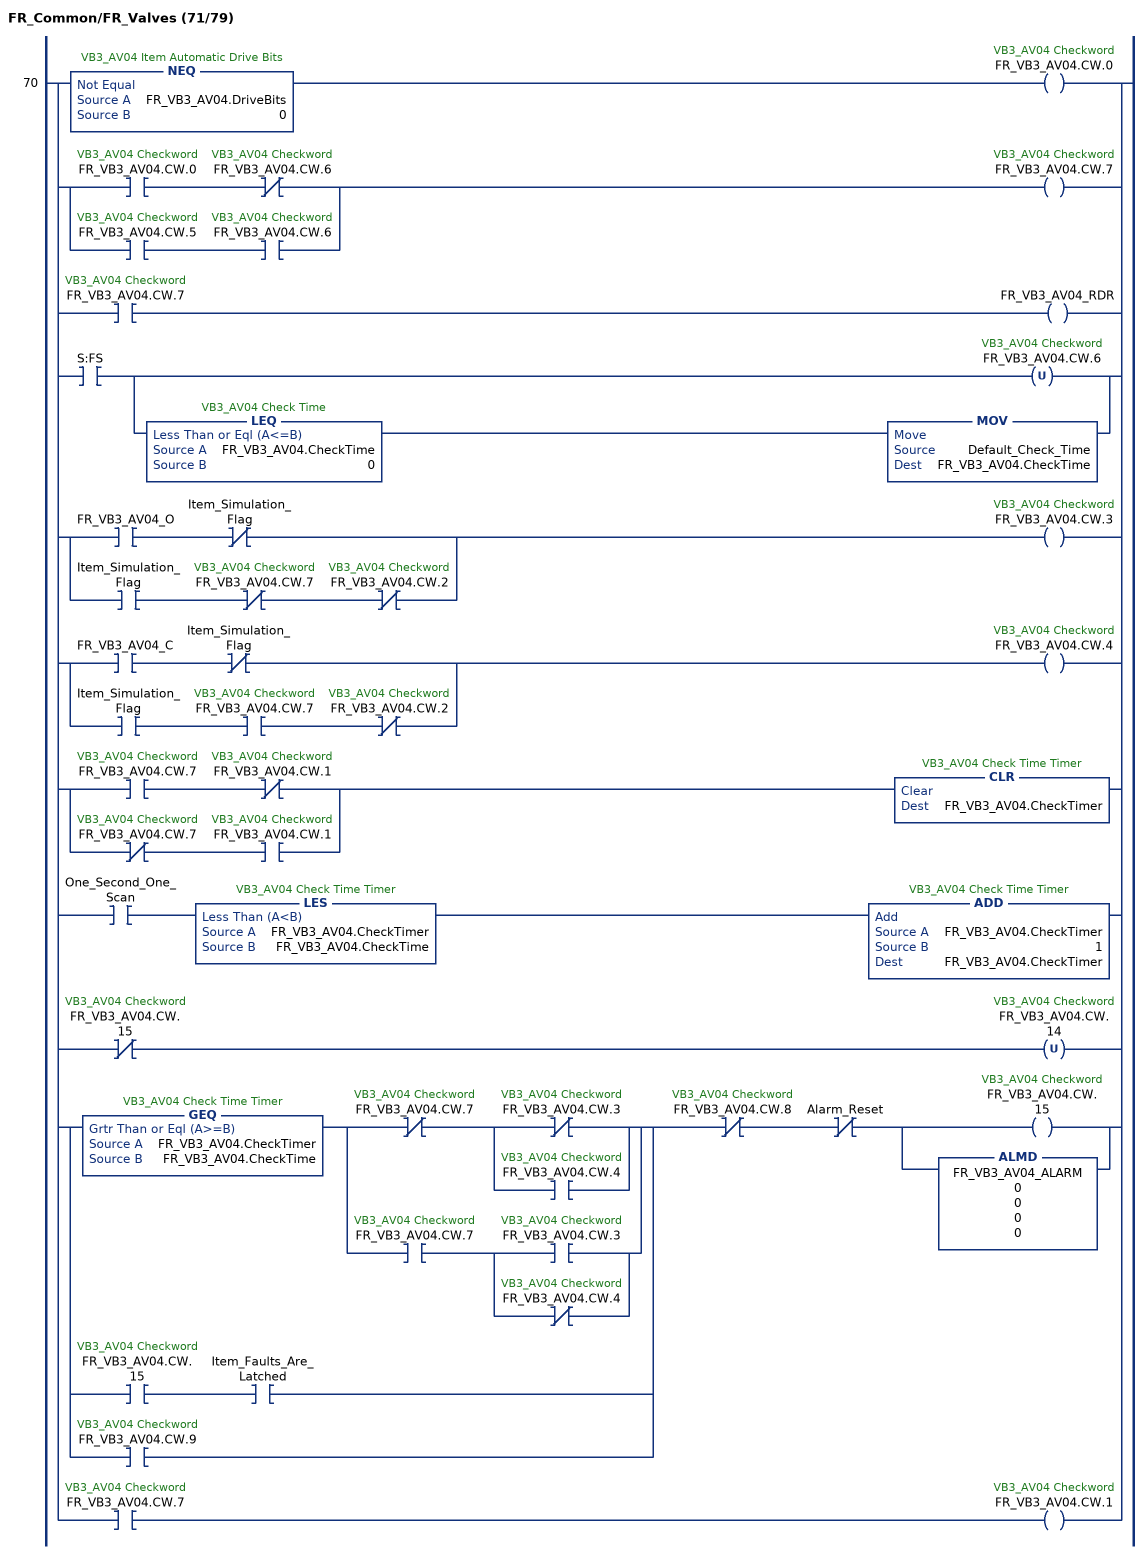
   70: [NEQ(FR_VB3_AV04.DriveBits,0) OTE(FR_VB3_AV04.CW.0) ,[XIC(FR_VB3_AV04.CW.0) XIO(FR_VB3_AV04.CW.6) ,XIC(FR_VB3_AV04.CW.5) XIC(FR_VB3_AV04.CW.6) ] OTE(FR_VB3_AV04.CW.7) ,XIC(FR_VB3_AV04.CW.7) OTE(FR_VB3_AV04_RDR) ,XIC(S:FS) [OTU(FR_VB3_AV04.CW.6) ,LEQ(FR_VB3_AV04.CheckTime,0) MOV(Default_Check_Time,FR_VB3_AV04.CheckTime) ] ,[[XIC(FR_VB3_AV04_O) XIO(Item_Simulation_Flag) ,XIC(Item_Simulation_Flag) XIO(FR_VB3_AV04.CW.7) XIO(FR_VB3_AV04.CW.2) ] OTE(FR_VB3_AV04.CW.3) ,[XIC(FR_VB3_AV04_C) XIO(Item_Simulation_Flag) ,XIC(Item_Simulation_Flag) XIC(FR_VB3_AV04.CW.7) XIO(FR_VB3_AV04.CW.2) ] OTE(FR_VB3_AV04.CW.4) ] ,[XIC(FR_VB3_AV04.CW.7) XIO(FR_VB3_AV04.CW.1) ,XIO(FR_VB3_AV04.CW.7) XIC(FR_VB3_AV04.CW.1) ] CLR(FR_VB3_AV04.CheckTimer) ,XIC(One_Second_One_Scan) LES(FR_VB3_AV04.CheckTimer,FR_VB3_AV04.CheckTime) ADD(FR_VB3_AV04.CheckTimer,1,FR_VB3_AV04.CheckTimer) ,XIO(FR_VB3_AV04.CW.15) OTU(FR_VB3_AV04.CW.14) ,[GEQ(FR_VB3_AV04.CheckTimer,FR_VB3_AV04.CheckTime) [XIO(FR_VB3_AV04.CW.7) [XIO(FR_VB3_AV04.CW.3) ,XIC(FR_VB3_AV04.CW.4) ] ,XIC(FR_VB3_AV04.CW.7) [XIC(FR_VB3_AV04.CW.3) ,XIO(FR_VB3_AV04.CW.4) ] ] ,XIC(FR_VB3_AV04.CW.15) XIC(Item_Faults_Are_Latched) ,XIC(FR_VB3_AV04.CW.9) ] XIO(FR_VB3_AV04.CW.8) XIO(Alarm_Reset) [OTE(FR_VB3_AV04.CW.15) ,ALMD(FR_VB3_AV04_ALARM,0,0,0,0) ] ,XIC(FR_VB3_AV04.CW.7) OTE(FR_VB3_AV04.CW.1) ];
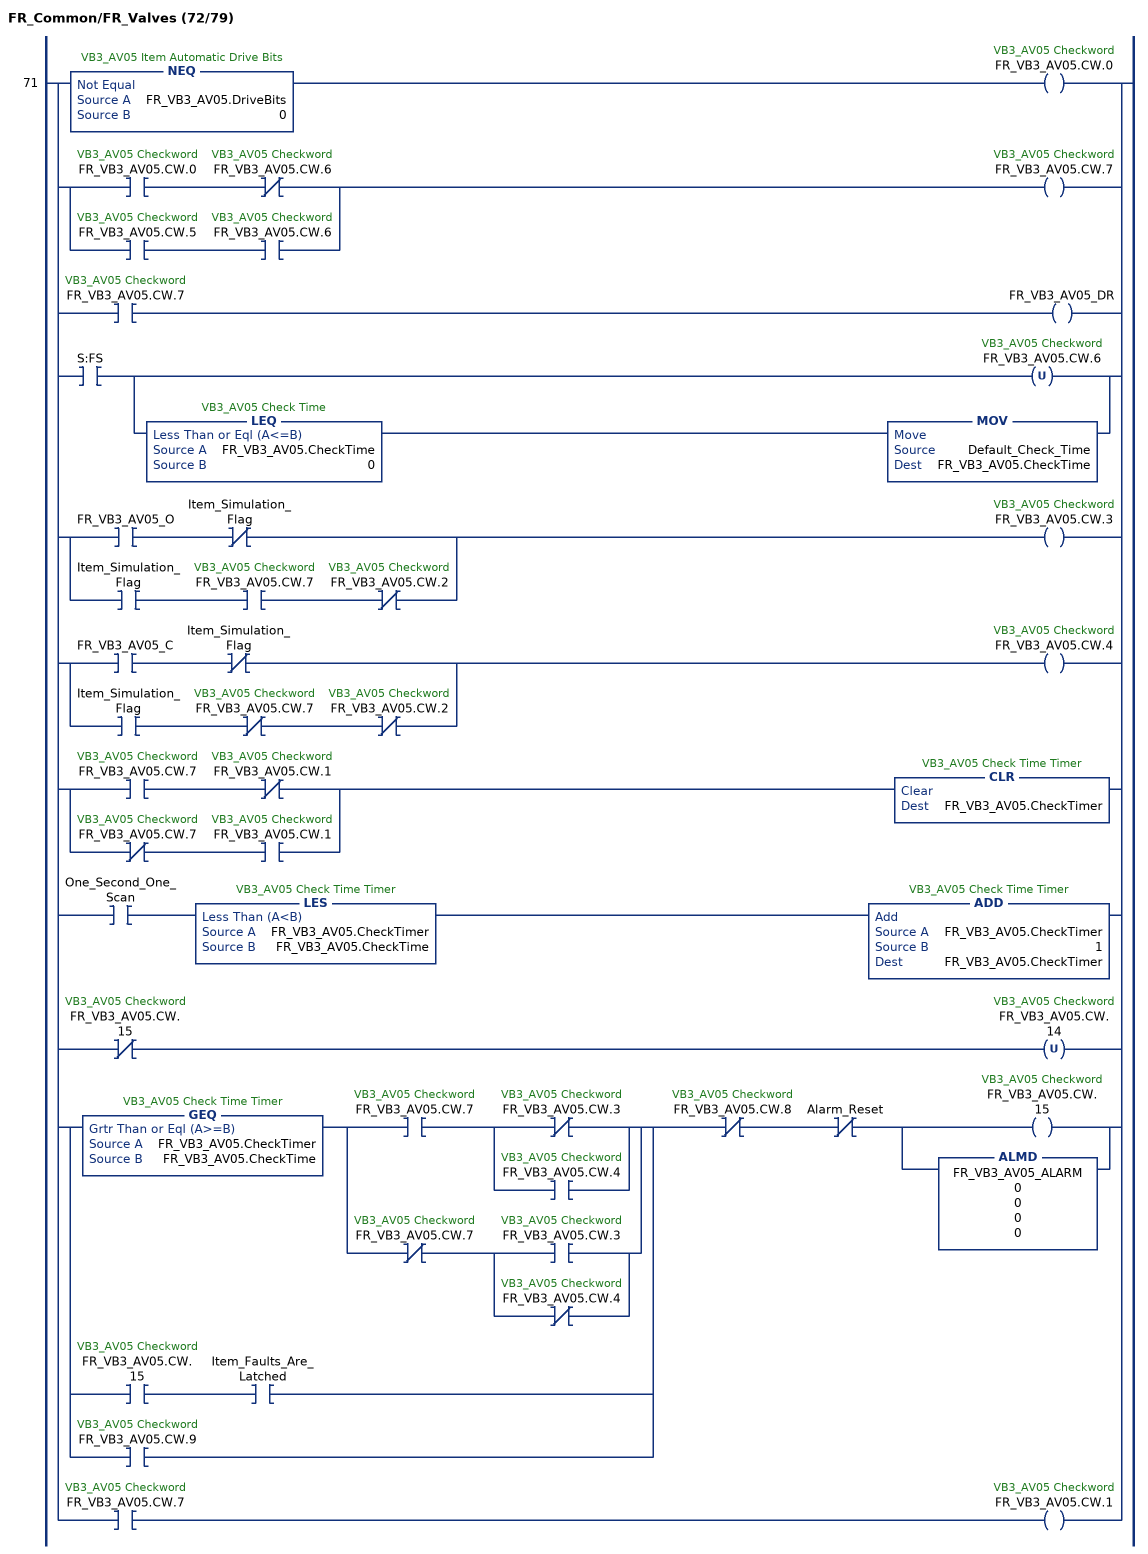
   71: [NEQ(FR_VB3_AV05.DriveBits,0) OTE(FR_VB3_AV05.CW.0) ,[XIC(FR_VB3_AV05.CW.0) XIO(FR_VB3_AV05.CW.6) ,XIC(FR_VB3_AV05.CW.5) XIC(FR_VB3_AV05.CW.6) ] OTE(FR_VB3_AV05.CW.7) ,XIC(FR_VB3_AV05.CW.7) OTE(FR_VB3_AV05_DR) ,XIC(S:FS) [OTU(FR_VB3_AV05.CW.6) ,LEQ(FR_VB3_AV05.CheckTime,0) MOV(Default_Check_Time,FR_VB3_AV05.CheckTime) ] ,[[XIC(FR_VB3_AV05_O) XIO(Item_Simulation_Flag) ,XIC(Item_Simulation_Flag) XIC(FR_VB3_AV05.CW.7) XIO(FR_VB3_AV05.CW.2) ] OTE(FR_VB3_AV05.CW.3) ,[XIC(FR_VB3_AV05_C) XIO(Item_Simulation_Flag) ,XIC(Item_Simulation_Flag) XIO(FR_VB3_AV05.CW.7) XIO(FR_VB3_AV05.CW.2) ] OTE(FR_VB3_AV05.CW.4) ] ,[XIC(FR_VB3_AV05.CW.7) XIO(FR_VB3_AV05.CW.1) ,XIO(FR_VB3_AV05.CW.7) XIC(FR_VB3_AV05.CW.1) ] CLR(FR_VB3_AV05.CheckTimer) ,XIC(One_Second_One_Scan) LES(FR_VB3_AV05.CheckTimer,FR_VB3_AV05.CheckTime) ADD(FR_VB3_AV05.CheckTimer,1,FR_VB3_AV05.CheckTimer) ,XIO(FR_VB3_AV05.CW.15) OTU(FR_VB3_AV05.CW.14) ,[GEQ(FR_VB3_AV05.CheckTimer,FR_VB3_AV05.CheckTime) [XIC(FR_VB3_AV05.CW.7) [XIO(FR_VB3_AV05.CW.3) ,XIC(FR_VB3_AV05.CW.4) ] ,XIO(FR_VB3_AV05.CW.7) [XIC(FR_VB3_AV05.CW.3) ,XIO(FR_VB3_AV05.CW.4) ] ] ,XIC(FR_VB3_AV05.CW.15) XIC(Item_Faults_Are_Latched) ,XIC(FR_VB3_AV05.CW.9) ] XIO(FR_VB3_AV05.CW.8) XIO(Alarm_Reset) [OTE(FR_VB3_AV05.CW.15) ,ALMD(FR_VB3_AV05_ALARM,0,0,0,0) ] ,XIC(FR_VB3_AV05.CW.7) OTE(FR_VB3_AV05.CW.1) ];
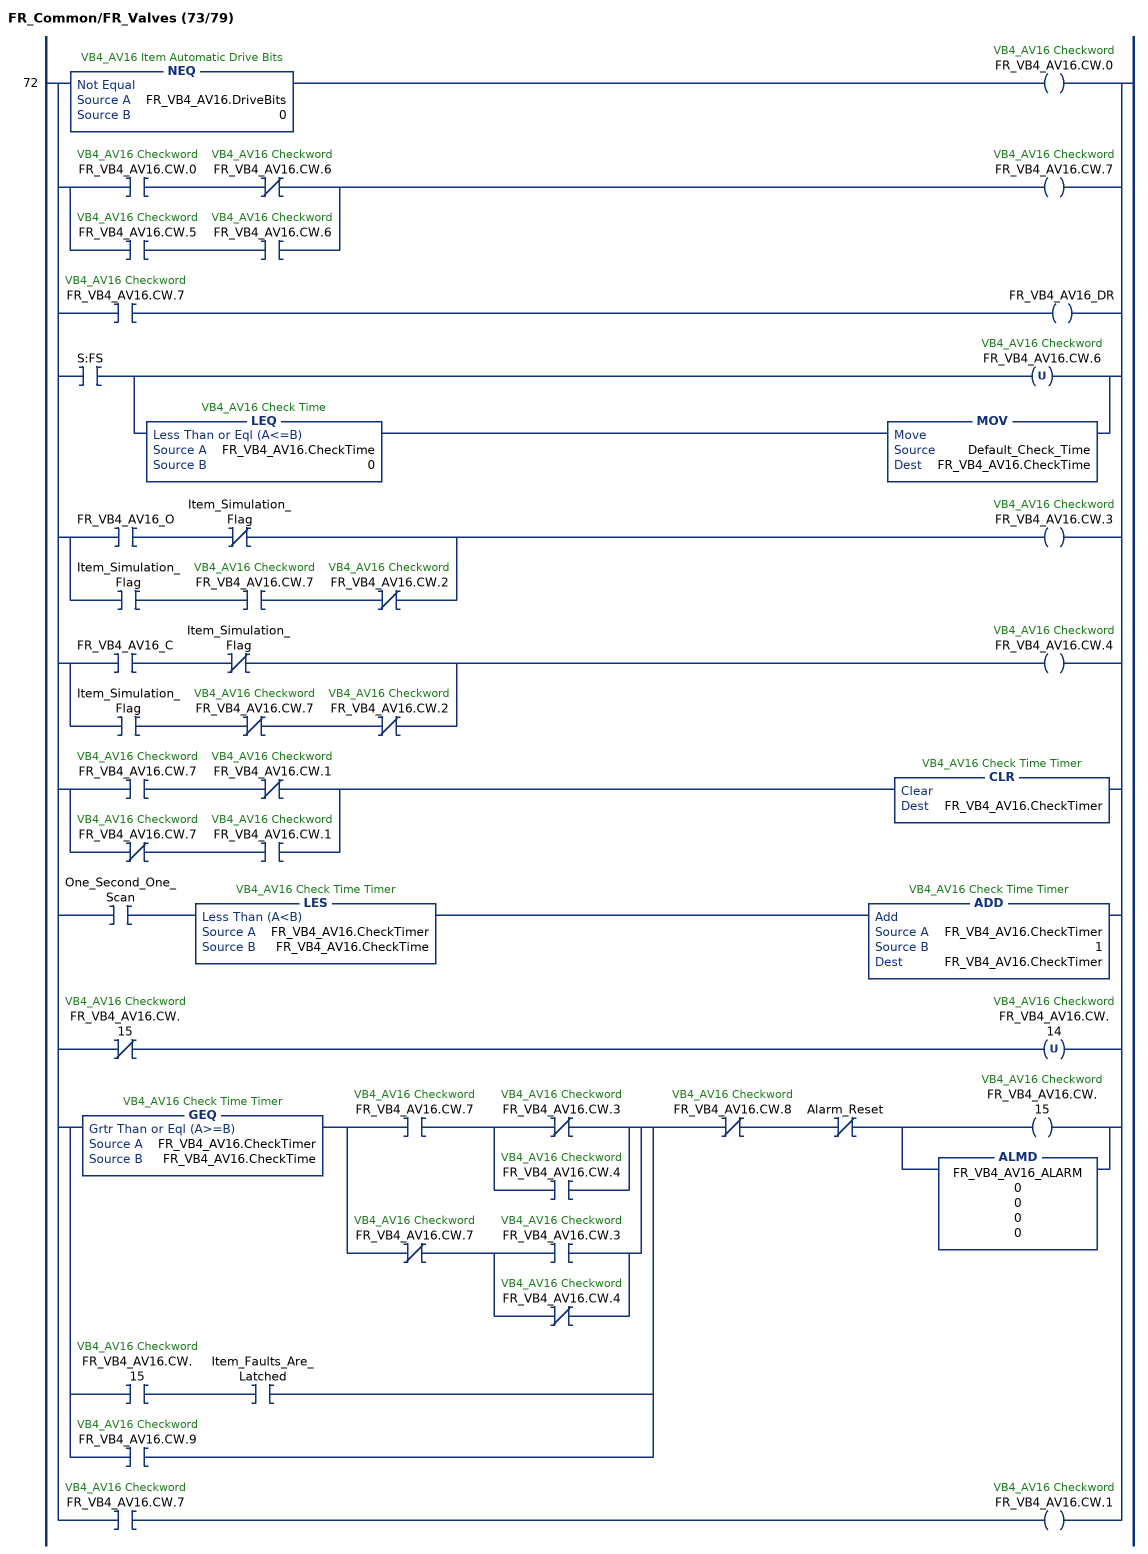
   72: [NEQ(FR_VB4_AV16.DriveBits,0) OTE(FR_VB4_AV16.CW.0) ,[XIC(FR_VB4_AV16.CW.0) XIO(FR_VB4_AV16.CW.6) ,XIC(FR_VB4_AV16.CW.5) XIC(FR_VB4_AV16.CW.6) ] OTE(FR_VB4_AV16.CW.7) ,XIC(FR_VB4_AV16.CW.7) OTE(FR_VB4_AV16_DR) ,XIC(S:FS) [OTU(FR_VB4_AV16.CW.6) ,LEQ(FR_VB4_AV16.CheckTime,0) MOV(Default_Check_Time,FR_VB4_AV16.CheckTime) ] ,[[XIC(FR_VB4_AV16_O) XIO(Item_Simulation_Flag) ,XIC(Item_Simulation_Flag) XIC(FR_VB4_AV16.CW.7) XIO(FR_VB4_AV16.CW.2) ] OTE(FR_VB4_AV16.CW.3) ,[XIC(FR_VB4_AV16_C) XIO(Item_Simulation_Flag) ,XIC(Item_Simulation_Flag) XIO(FR_VB4_AV16.CW.7) XIO(FR_VB4_AV16.CW.2) ] OTE(FR_VB4_AV16.CW.4) ] ,[XIC(FR_VB4_AV16.CW.7) XIO(FR_VB4_AV16.CW.1) ,XIO(FR_VB4_AV16.CW.7) XIC(FR_VB4_AV16.CW.1) ] CLR(FR_VB4_AV16.CheckTimer) ,XIC(One_Second_One_Scan) LES(FR_VB4_AV16.CheckTimer,FR_VB4_AV16.CheckTime) ADD(FR_VB4_AV16.CheckTimer,1,FR_VB4_AV16.CheckTimer) ,XIO(FR_VB4_AV16.CW.15) OTU(FR_VB4_AV16.CW.14) ,[GEQ(FR_VB4_AV16.CheckTimer,FR_VB4_AV16.CheckTime) [XIC(FR_VB4_AV16.CW.7) [XIO(FR_VB4_AV16.CW.3) ,XIC(FR_VB4_AV16.CW.4) ] ,XIO(FR_VB4_AV16.CW.7) [XIC(FR_VB4_AV16.CW.3) ,XIO(FR_VB4_AV16.CW.4) ] ] ,XIC(FR_VB4_AV16.CW.15) XIC(Item_Faults_Are_Latched) ,XIC(FR_VB4_AV16.CW.9) ] XIO(FR_VB4_AV16.CW.8) XIO(Alarm_Reset) [OTE(FR_VB4_AV16.CW.15) ,ALMD(FR_VB4_AV16_ALARM,0,0,0,0) ] ,XIC(FR_VB4_AV16.CW.7) OTE(FR_VB4_AV16.CW.1) ];
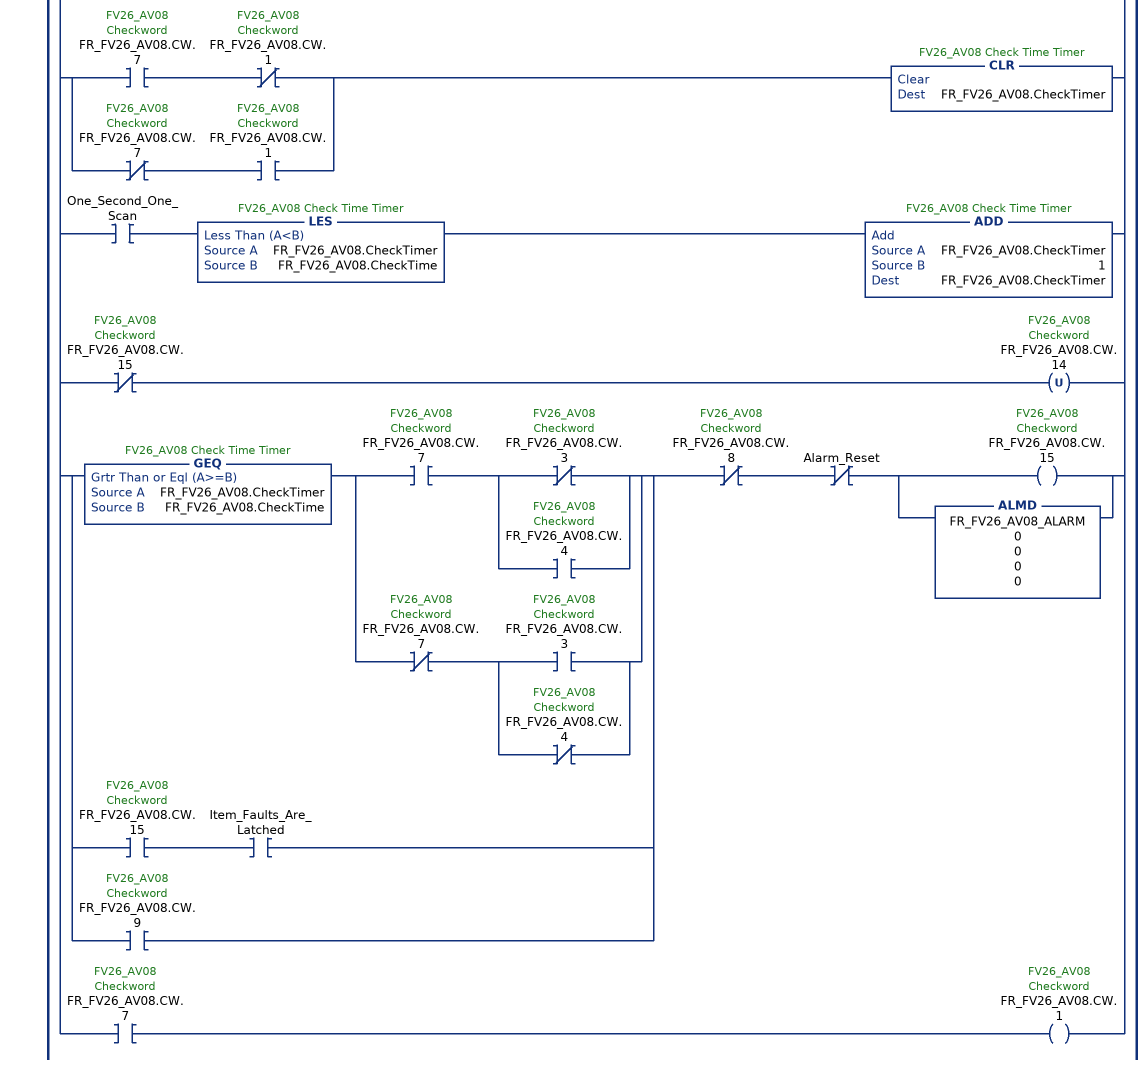
   73: [NEQ(FR_FV26_AV08.DriveBits,0) OTE(FR_FV26_AV08.CW.0) ,[XIC(FR_FV26_AV08.CW.0) XIO(FR_FV26_AV08.CW.6) ,XIC(FR_FV26_AV08.CW.5) XIC(FR_FV26_AV08.CW.6) ] OTE(FR_FV26_AV08.CW.7) ,XIC(FR_FV26_AV08.CW.7) OTE(FR_FV26_AV08_DR) ,XIC(S:FS) [OTU(FR_FV26_AV08.CW.6) ,LEQ(FR_FV26_AV08.CheckTime,0) MOV(Default_Check_Time,FR_FV26_AV08.CheckTime) ] ,[[XIC(FR_FV26_AV08_O) XIO(Item_Simulation_Flag) ,XIC(Item_Simulation_Flag) XIC(FR_FV26_AV08.CW.7) XIO(FR_FV26_AV08.CW.2) ] OTE(FR_FV26_AV08.CW.3) ,[XIC(FR_FV26_AV08_C) XIO(Item_Simulation_Flag) ,XIC(Item_Simulation_Flag) XIO(FR_FV26_AV08.CW.7) XIO(FR_FV26_AV08.CW.2) ] OTE(FR_FV26_AV08.CW.4) ] ,[XIC(FR_FV26_AV08.CW.7) XIO(FR_FV26_AV08.CW.1) ,XIO(FR_FV26_AV08.CW.7) XIC(FR_FV26_AV08.CW.1) ] CLR(FR_FV26_AV08.CheckTimer) ,XIC(One_Second_One_Scan) LES(FR_FV26_AV08.CheckTimer,FR_FV26_AV08.CheckTime) ADD(FR_FV26_AV08.CheckTimer,1,FR_FV26_AV08.CheckTimer) ,XIO(FR_FV26_AV08.CW.15) OTU(FR_FV26_AV08.CW.14) ,[GEQ(FR_FV26_AV08.CheckTimer,FR_FV26_AV08.CheckTime) [XIC(FR_FV26_AV08.CW.7) [XIO(FR_FV26_AV08.CW.3) ,XIC(FR_FV26_AV08.CW.4) ] ,XIO(FR_FV26_AV08.CW.7) [XIC(FR_FV26_AV08.CW.3) ,XIO(FR_FV26_AV08.CW.4) ] ] ,XIC(FR_FV26_AV08.CW.15) XIC(Item_Faults_Are_Latched) ,XIC(FR_FV26_AV08.CW.9) ] XIO(FR_FV26_AV08.CW.8) XIO(Alarm_Reset) [OTE(FR_FV26_AV08.CW.15) ,ALMD(FR_FV26_AV08_ALARM,0,0,0,0) ] ,XIC(FR_FV26_AV08.CW.7) OTE(FR_FV26_AV08.CW.1) ];
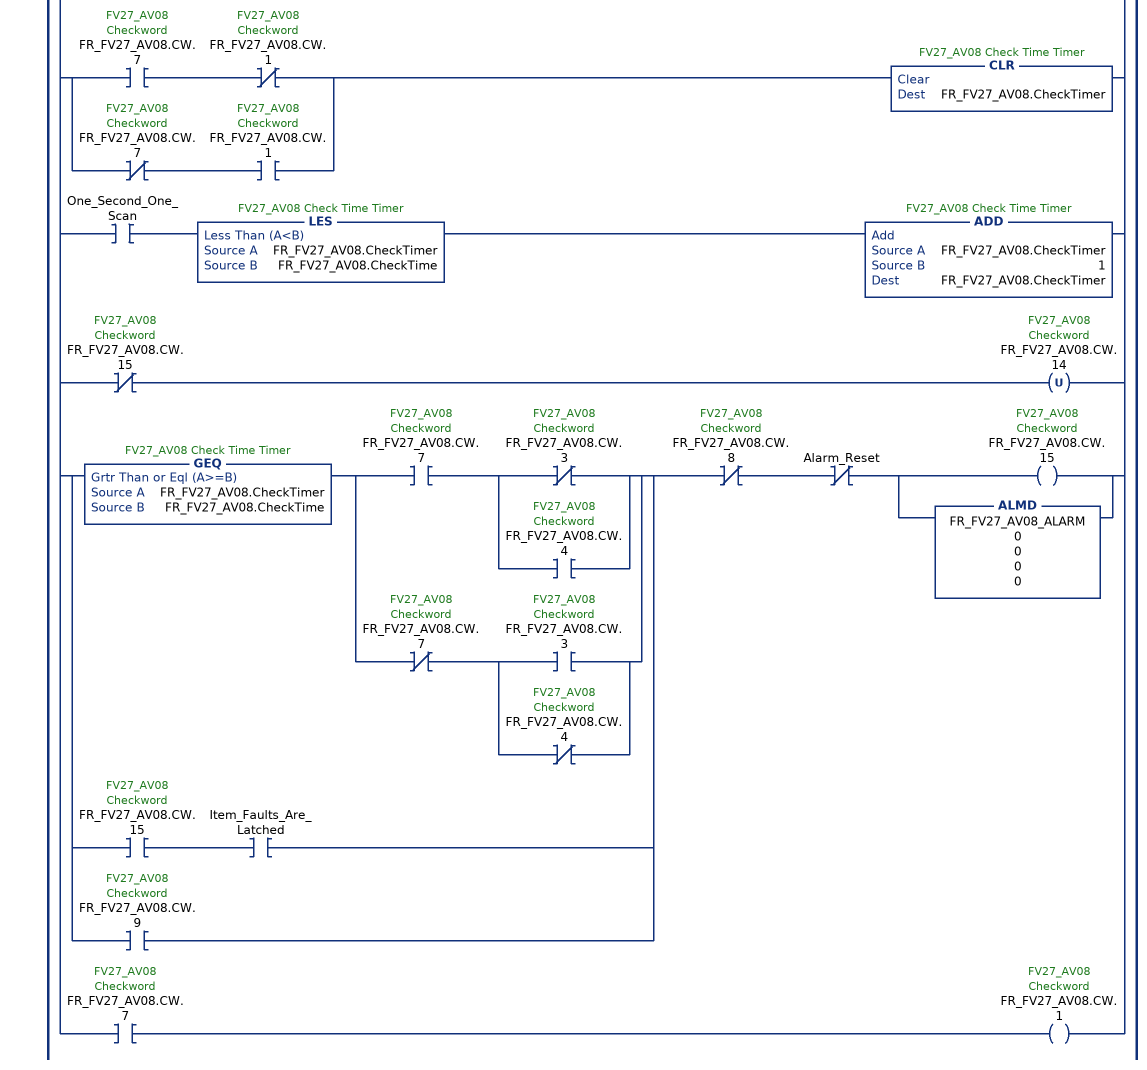
   74: [NEQ(FR_FV27_AV08.DriveBits,0) OTE(FR_FV27_AV08.CW.0) ,[XIC(FR_FV27_AV08.CW.0) XIO(FR_FV27_AV08.CW.6) ,XIC(FR_FV27_AV08.CW.5) XIC(FR_FV27_AV08.CW.6) ] OTE(FR_FV27_AV08.CW.7) ,XIC(FR_FV27_AV08.CW.7) OTE(FR_FV27_AV08_DR) ,XIC(S:FS) [OTU(FR_FV27_AV08.CW.6) ,LEQ(FR_FV27_AV08.CheckTime,0) MOV(Default_Check_Time,FR_FV27_AV08.CheckTime) ] ,[[XIC(FR_FV27_AV08_O) XIO(Item_Simulation_Flag) ,XIC(Item_Simulation_Flag) XIC(FR_FV27_AV08.CW.7) XIO(FR_FV27_AV08.CW.2) ] OTE(FR_FV27_AV08.CW.3) ,[XIC(FR_FV27_AV08_C) XIO(Item_Simulation_Flag) ,XIC(Item_Simulation_Flag) XIO(FR_FV27_AV08.CW.7) XIO(FR_FV27_AV08.CW.2) ] OTE(FR_FV27_AV08.CW.4) ] ,[XIC(FR_FV27_AV08.CW.7) XIO(FR_FV27_AV08.CW.1) ,XIO(FR_FV27_AV08.CW.7) XIC(FR_FV27_AV08.CW.1) ] CLR(FR_FV27_AV08.CheckTimer) ,XIC(One_Second_One_Scan) LES(FR_FV27_AV08.CheckTimer,FR_FV27_AV08.CheckTime) ADD(FR_FV27_AV08.CheckTimer,1,FR_FV27_AV08.CheckTimer) ,XIO(FR_FV27_AV08.CW.15) OTU(FR_FV27_AV08.CW.14) ,[GEQ(FR_FV27_AV08.CheckTimer,FR_FV27_AV08.CheckTime) [XIC(FR_FV27_AV08.CW.7) [XIO(FR_FV27_AV08.CW.3) ,XIC(FR_FV27_AV08.CW.4) ] ,XIO(FR_FV27_AV08.CW.7) [XIC(FR_FV27_AV08.CW.3) ,XIO(FR_FV27_AV08.CW.4) ] ] ,XIC(FR_FV27_AV08.CW.15) XIC(Item_Faults_Are_Latched) ,XIC(FR_FV27_AV08.CW.9) ] XIO(FR_FV27_AV08.CW.8) XIO(Alarm_Reset) [OTE(FR_FV27_AV08.CW.15) ,ALMD(FR_FV27_AV08_ALARM,0,0,0,0) ] ,XIC(FR_FV27_AV08.CW.7) OTE(FR_FV27_AV08.CW.1) ];
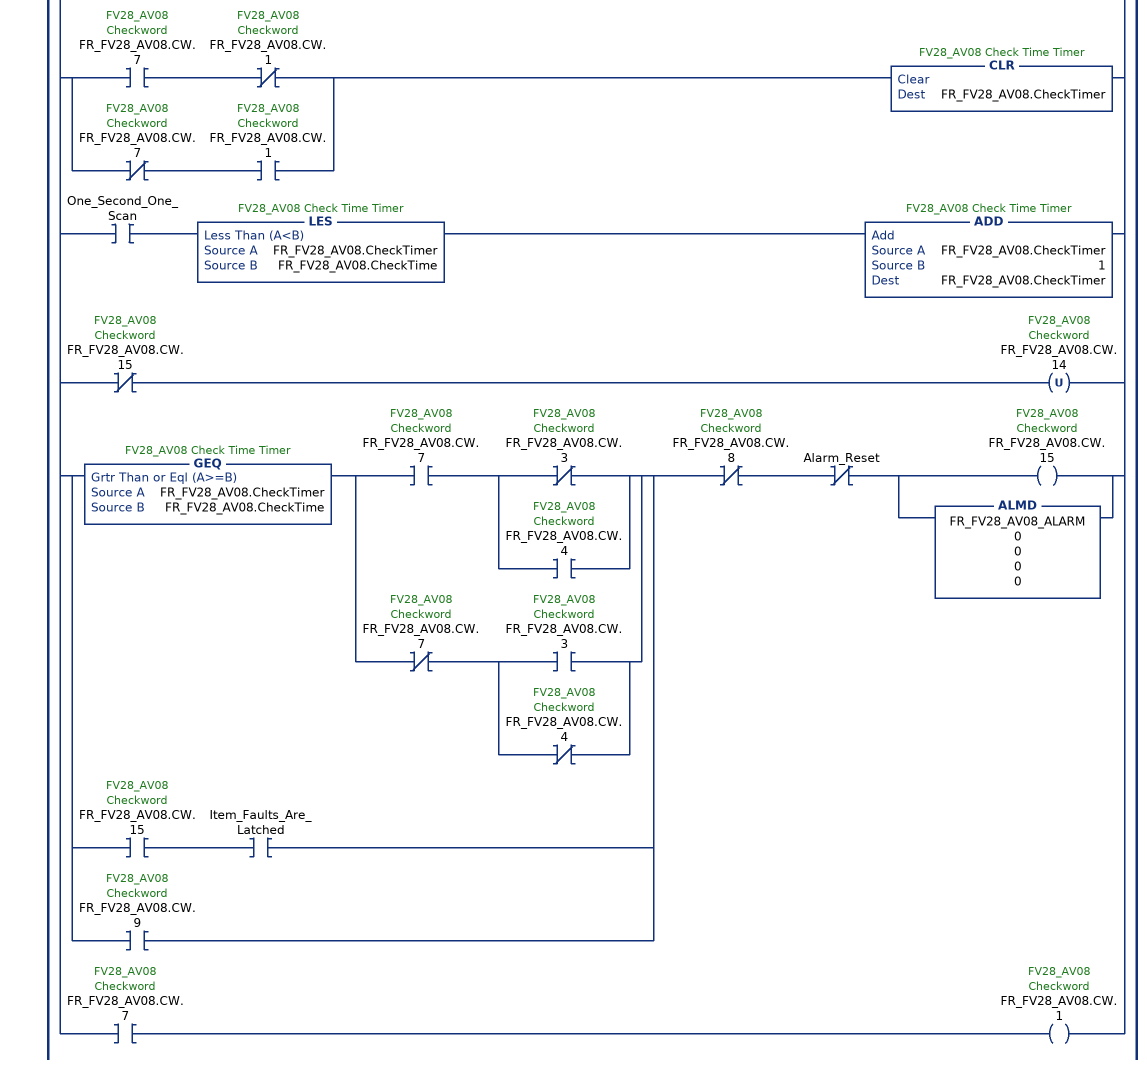
   75: [NEQ(FR_FV28_AV08.DriveBits,0) OTE(FR_FV28_AV08.CW.0) ,[XIC(FR_FV28_AV08.CW.0) XIO(FR_FV28_AV08.CW.6) ,XIC(FR_FV28_AV08.CW.5) XIC(FR_FV28_AV08.CW.6) ] OTE(FR_FV28_AV08.CW.7) ,XIC(FR_FV28_AV08.CW.7) OTE(FR_FV28_AV08_DR) ,XIC(S:FS) [OTU(FR_FV28_AV08.CW.6) ,LEQ(FR_FV28_AV08.CheckTime,0) MOV(Default_Check_Time,FR_FV28_AV08.CheckTime) ] ,[[XIC(FR_FV28_AV08_O) XIO(Item_Simulation_Flag) ,XIC(Item_Simulation_Flag) XIC(FR_FV28_AV08.CW.7) XIO(FR_FV28_AV08.CW.2) ] OTE(FR_FV28_AV08.CW.3) ,[XIC(FR_FV28_AV08_C) XIO(Item_Simulation_Flag) ,XIC(Item_Simulation_Flag) XIO(FR_FV28_AV08.CW.7) XIO(FR_FV28_AV08.CW.2) ] OTE(FR_FV28_AV08.CW.4) ] ,[XIC(FR_FV28_AV08.CW.7) XIO(FR_FV28_AV08.CW.1) ,XIO(FR_FV28_AV08.CW.7) XIC(FR_FV28_AV08.CW.1) ] CLR(FR_FV28_AV08.CheckTimer) ,XIC(One_Second_One_Scan) LES(FR_FV28_AV08.CheckTimer,FR_FV28_AV08.CheckTime) ADD(FR_FV28_AV08.CheckTimer,1,FR_FV28_AV08.CheckTimer) ,XIO(FR_FV28_AV08.CW.15) OTU(FR_FV28_AV08.CW.14) ,[GEQ(FR_FV28_AV08.CheckTimer,FR_FV28_AV08.CheckTime) [XIC(FR_FV28_AV08.CW.7) [XIO(FR_FV28_AV08.CW.3) ,XIC(FR_FV28_AV08.CW.4) ] ,XIO(FR_FV28_AV08.CW.7) [XIC(FR_FV28_AV08.CW.3) ,XIO(FR_FV28_AV08.CW.4) ] ] ,XIC(FR_FV28_AV08.CW.15) XIC(Item_Faults_Are_Latched) ,XIC(FR_FV28_AV08.CW.9) ] XIO(FR_FV28_AV08.CW.8) XIO(Alarm_Reset) [OTE(FR_FV28_AV08.CW.15) ,ALMD(FR_FV28_AV08_ALARM,0,0,0,0) ] ,XIC(FR_FV28_AV08.CW.7) OTE(FR_FV28_AV08.CW.1) ];
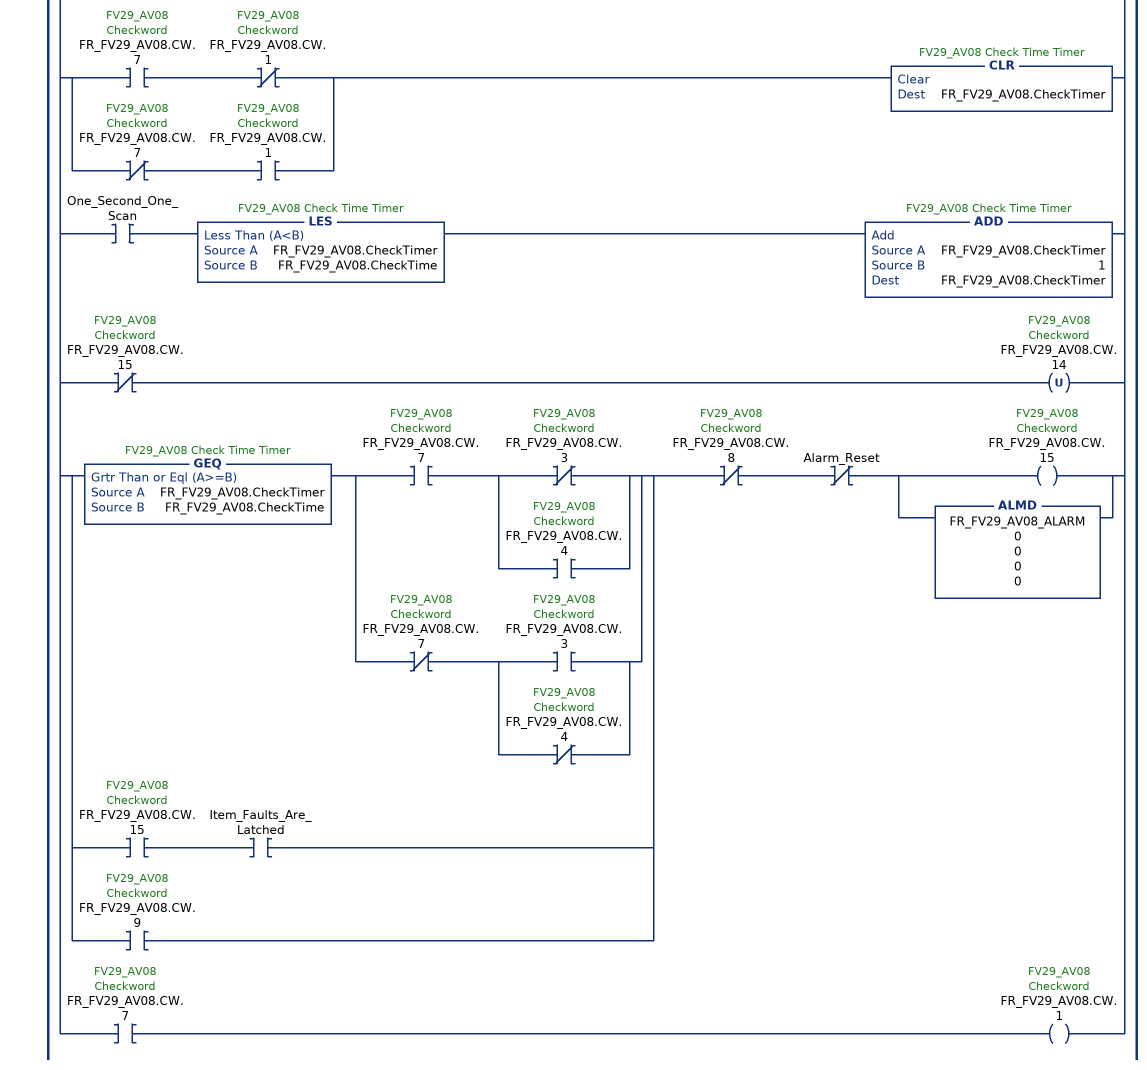
   76: [NEQ(FR_FV29_AV08.DriveBits,0) OTE(FR_FV29_AV08.CW.0) ,[XIC(FR_FV29_AV08.CW.0) XIO(FR_FV29_AV08.CW.6) ,XIC(FR_FV29_AV08.CW.5) XIC(FR_FV29_AV08.CW.6) ] OTE(FR_FV29_AV08.CW.7) ,XIC(FR_FV29_AV08.CW.7) OTE(FR_FV29_AV08_DR) ,XIC(S:FS) [OTU(FR_FV29_AV08.CW.6) ,LEQ(FR_FV29_AV08.CheckTime,0) MOV(Default_Check_Time,FR_FV29_AV08.CheckTime) ] ,[[XIC(FR_FV29_AV08_O) XIO(Item_Simulation_Flag) ,XIC(Item_Simulation_Flag) XIC(FR_FV29_AV08.CW.7) XIO(FR_FV29_AV08.CW.2) ] OTE(FR_FV29_AV08.CW.3) ,[XIC(FR_FV29_AV08_C) XIO(Item_Simulation_Flag) ,XIC(Item_Simulation_Flag) XIO(FR_FV29_AV08.CW.7) XIO(FR_FV29_AV08.CW.2) ] OTE(FR_FV29_AV08.CW.4) ] ,[XIC(FR_FV29_AV08.CW.7) XIO(FR_FV29_AV08.CW.1) ,XIO(FR_FV29_AV08.CW.7) XIC(FR_FV29_AV08.CW.1) ] CLR(FR_FV29_AV08.CheckTimer) ,XIC(One_Second_One_Scan) LES(FR_FV29_AV08.CheckTimer,FR_FV29_AV08.CheckTime) ADD(FR_FV29_AV08.CheckTimer,1,FR_FV29_AV08.CheckTimer) ,XIO(FR_FV29_AV08.CW.15) OTU(FR_FV29_AV08.CW.14) ,[GEQ(FR_FV29_AV08.CheckTimer,FR_FV29_AV08.CheckTime) [XIC(FR_FV29_AV08.CW.7) [XIO(FR_FV29_AV08.CW.3) ,XIC(FR_FV29_AV08.CW.4) ] ,XIO(FR_FV29_AV08.CW.7) [XIC(FR_FV29_AV08.CW.3) ,XIO(FR_FV29_AV08.CW.4) ] ] ,XIC(FR_FV29_AV08.CW.15) XIC(Item_Faults_Are_Latched) ,XIC(FR_FV29_AV08.CW.9) ] XIO(FR_FV29_AV08.CW.8) XIO(Alarm_Reset) [OTE(FR_FV29_AV08.CW.15) ,ALMD(FR_FV29_AV08_ALARM,0,0,0,0) ] ,XIC(FR_FV29_AV08.CW.7) OTE(FR_FV29_AV08.CW.1) ];
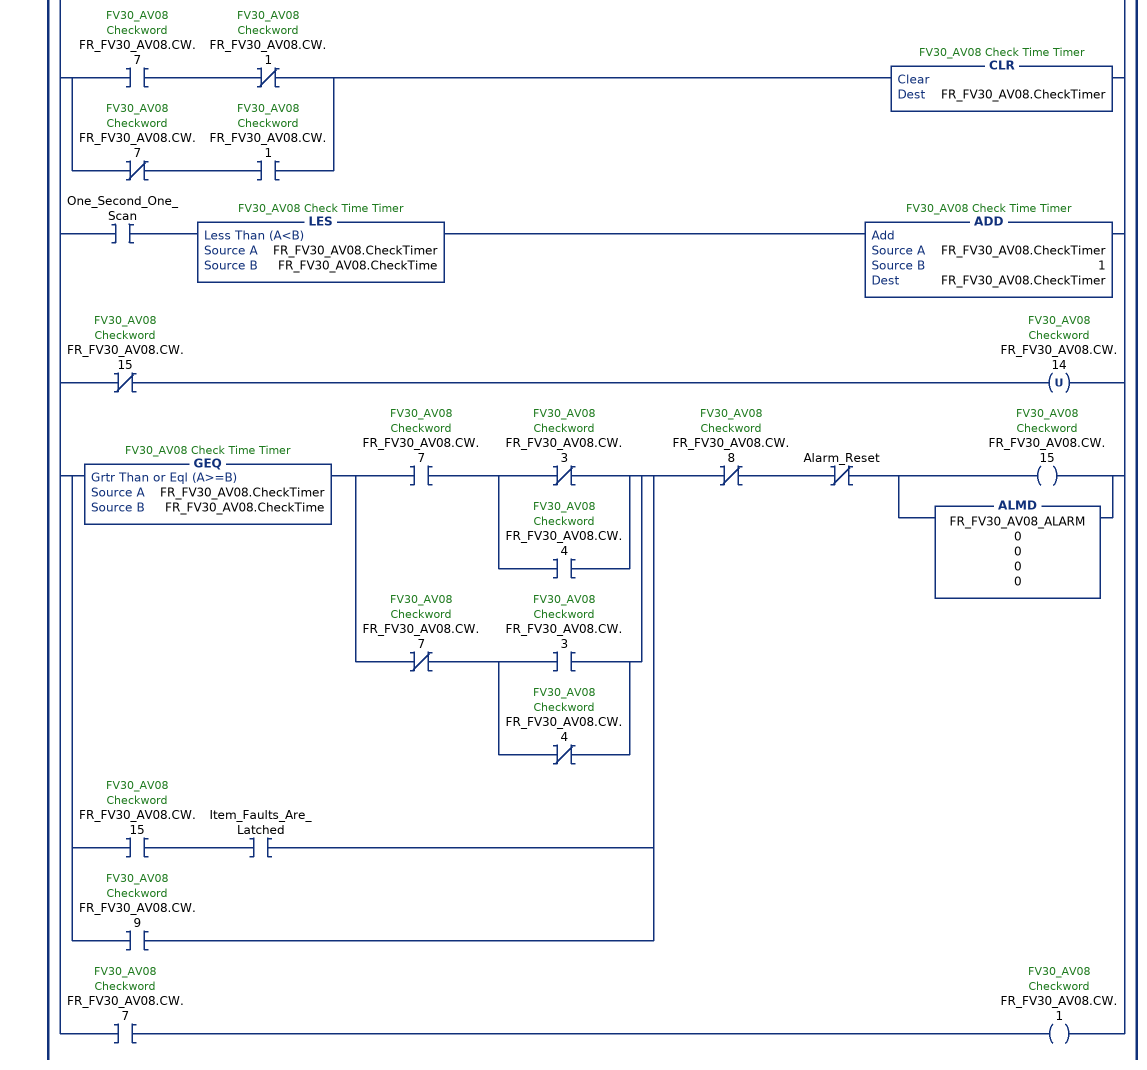
   77: [NEQ(FR_FV30_AV08.DriveBits,0) OTE(FR_FV30_AV08.CW.0) ,[XIC(FR_FV30_AV08.CW.0) XIO(FR_FV30_AV08.CW.6) ,XIC(FR_FV30_AV08.CW.5) XIC(FR_FV30_AV08.CW.6) ] OTE(FR_FV30_AV08.CW.7) ,XIC(FR_FV30_AV08.CW.7) OTE(FR_FV30_AV08_DR) ,XIC(S:FS) [OTU(FR_FV30_AV08.CW.6) ,LEQ(FR_FV30_AV08.CheckTime,0) MOV(Default_Check_Time,FR_FV30_AV08.CheckTime) ] ,[[XIC(FR_FV30_AV08_O) XIO(Item_Simulation_Flag) ,XIC(Item_Simulation_Flag) XIC(FR_FV30_AV08.CW.7) XIO(FR_FV30_AV08.CW.2) ] OTE(FR_FV30_AV08.CW.3) ,[XIC(FR_FV30_AV08_C) XIO(Item_Simulation_Flag) ,XIC(Item_Simulation_Flag) XIO(FR_FV30_AV08.CW.7) XIO(FR_FV30_AV08.CW.2) ] OTE(FR_FV30_AV08.CW.4) ] ,[XIC(FR_FV30_AV08.CW.7) XIO(FR_FV30_AV08.CW.1) ,XIO(FR_FV30_AV08.CW.7) XIC(FR_FV30_AV08.CW.1) ] CLR(FR_FV30_AV08.CheckTimer) ,XIC(One_Second_One_Scan) LES(FR_FV30_AV08.CheckTimer,FR_FV30_AV08.CheckTime) ADD(FR_FV30_AV08.CheckTimer,1,FR_FV30_AV08.CheckTimer) ,XIO(FR_FV30_AV08.CW.15) OTU(FR_FV30_AV08.CW.14) ,[GEQ(FR_FV30_AV08.CheckTimer,FR_FV30_AV08.CheckTime) [XIC(FR_FV30_AV08.CW.7) [XIO(FR_FV30_AV08.CW.3) ,XIC(FR_FV30_AV08.CW.4) ] ,XIO(FR_FV30_AV08.CW.7) [XIC(FR_FV30_AV08.CW.3) ,XIO(FR_FV30_AV08.CW.4) ] ] ,XIC(FR_FV30_AV08.CW.15) XIC(Item_Faults_Are_Latched) ,XIC(FR_FV30_AV08.CW.9) ] XIO(FR_FV30_AV08.CW.8) XIO(Alarm_Reset) [OTE(FR_FV30_AV08.CW.15) ,ALMD(FR_FV30_AV08_ALARM,0,0,0,0) ] ,XIC(FR_FV30_AV08.CW.7) OTE(FR_FV30_AV08.CW.1) ];
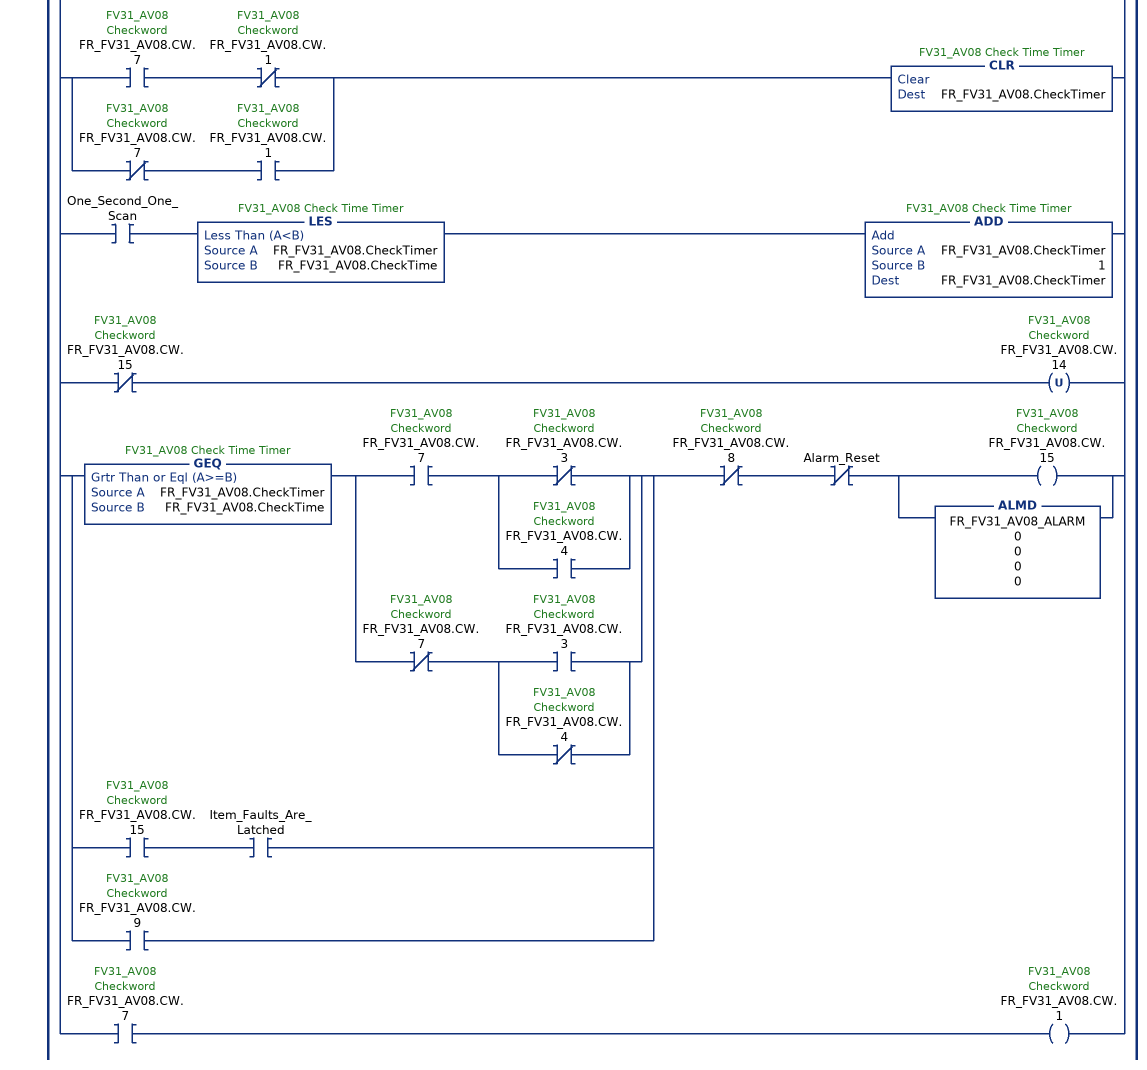
   78: [NEQ(FR_FV31_AV08.DriveBits,0) OTE(FR_FV31_AV08.CW.0) ,[XIC(FR_FV31_AV08.CW.0) XIO(FR_FV31_AV08.CW.6) ,XIC(FR_FV31_AV08.CW.5) XIC(FR_FV31_AV08.CW.6) ] OTE(FR_FV31_AV08.CW.7) ,XIC(FR_FV31_AV08.CW.7) OTE(FR_FV31_AV08_DR) ,XIC(S:FS) [OTU(FR_FV31_AV08.CW.6) ,LEQ(FR_FV31_AV08.CheckTime,0) MOV(Default_Check_Time,FR_FV31_AV08.CheckTime) ] ,[[[XIC(FR_FV31_AV08_O) ,XIC(FR_FV31_AV08_O1) ] XIO(Item_Simulation_Flag) ,XIC(Item_Simulation_Flag) XIC(FR_FV31_AV08.CW.7) XIO(FR_FV31_AV08.CW.2) ] OTE(FR_FV31_AV08.CW.3) ,[XIC(FR_FV31_AV08_C) XIO(Item_Simulation_Flag) ,XIC(Item_Simulation_Flag) XIO(FR_FV31_AV08.CW.7) XIO(FR_FV31_AV08.CW.2) ] OTE(FR_FV31_AV08.CW.4) ] ,[XIC(FR_FV31_AV08.CW.7) XIO(FR_FV31_AV08.CW.1) ,XIO(FR_FV31_AV08.CW.7) XIC(FR_FV31_AV08.CW.1) ] CLR(FR_FV31_AV08.CheckTimer) ,XIC(One_Second_One_Scan) LES(FR_FV31_AV08.CheckTimer,FR_FV31_AV08.CheckTime) ADD(FR_FV31_AV08.CheckTimer,1,FR_FV31_AV08.CheckTimer) ,XIO(FR_FV31_AV08.CW.15) OTU(FR_FV31_AV08.CW.14) ,[GEQ(FR_FV31_AV08.CheckTimer,FR_FV31_AV08.CheckTime) [XIC(FR_FV31_AV08.CW.7) [XIO(FR_FV31_AV08.CW.3) ,XIC(FR_FV31_AV08.CW.4) ] ,XIO(FR_FV31_AV08.CW.7) [XIC(FR_FV31_AV08.CW.3) ,XIO(FR_FV31_AV08.CW.4) ] ] ,XIC(FR_FV31_AV08.CW.15) XIC(Item_Faults_Are_Latched) ,XIC(FR_FV31_AV08.CW.9) ] XIO(FR_FV31_AV08.CW.8) XIO(Alarm_Reset) [OTE(FR_FV31_AV08.CW.15) ,ALMD(FR_FV31_AV08_ALARM,0,0,0,0) ] ,XIC(FR_FV31_AV08.CW.7) OTE(FR_FV31_AV08.CW.1) ];
END_ROUTINE

ROUTINE FR_Vent_Drives   (* ladder *)
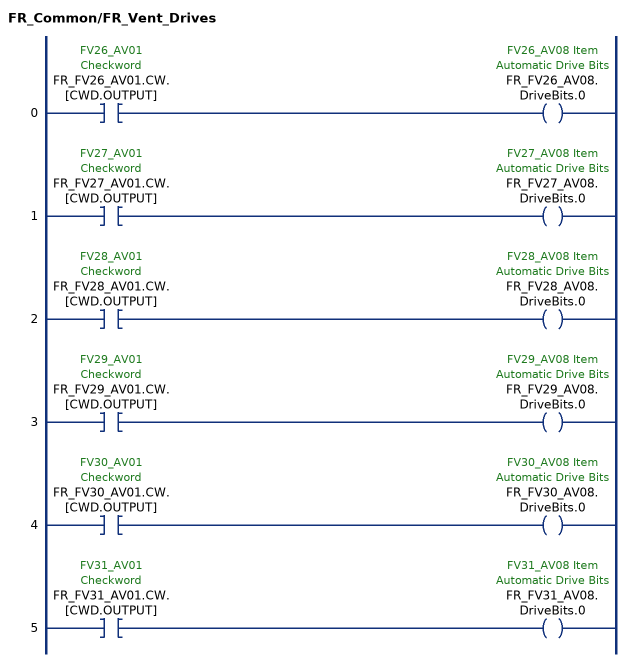
   0: XIC(FR_FV26_AV01.CW.[CWD.OUTPUT])OTE(FR_FV26_AV08.DriveBits.0);
   1: XIC(FR_FV27_AV01.CW.[CWD.OUTPUT])OTE(FR_FV27_AV08.DriveBits.0);
   2: XIC(FR_FV28_AV01.CW.[CWD.OUTPUT])OTE(FR_FV28_AV08.DriveBits.0);
   3: XIC(FR_FV29_AV01.CW.[CWD.OUTPUT])OTE(FR_FV29_AV08.DriveBits.0);
   4: XIC(FR_FV30_AV01.CW.[CWD.OUTPUT])OTE(FR_FV30_AV08.DriveBits.0);
   5: XIC(FR_FV31_AV01.CW.[CWD.OUTPUT])OTE(FR_FV31_AV08.DriveBits.0);
END_ROUTINE
